// TIA Portal project "DistributoreCaffè" (V19) (continued)
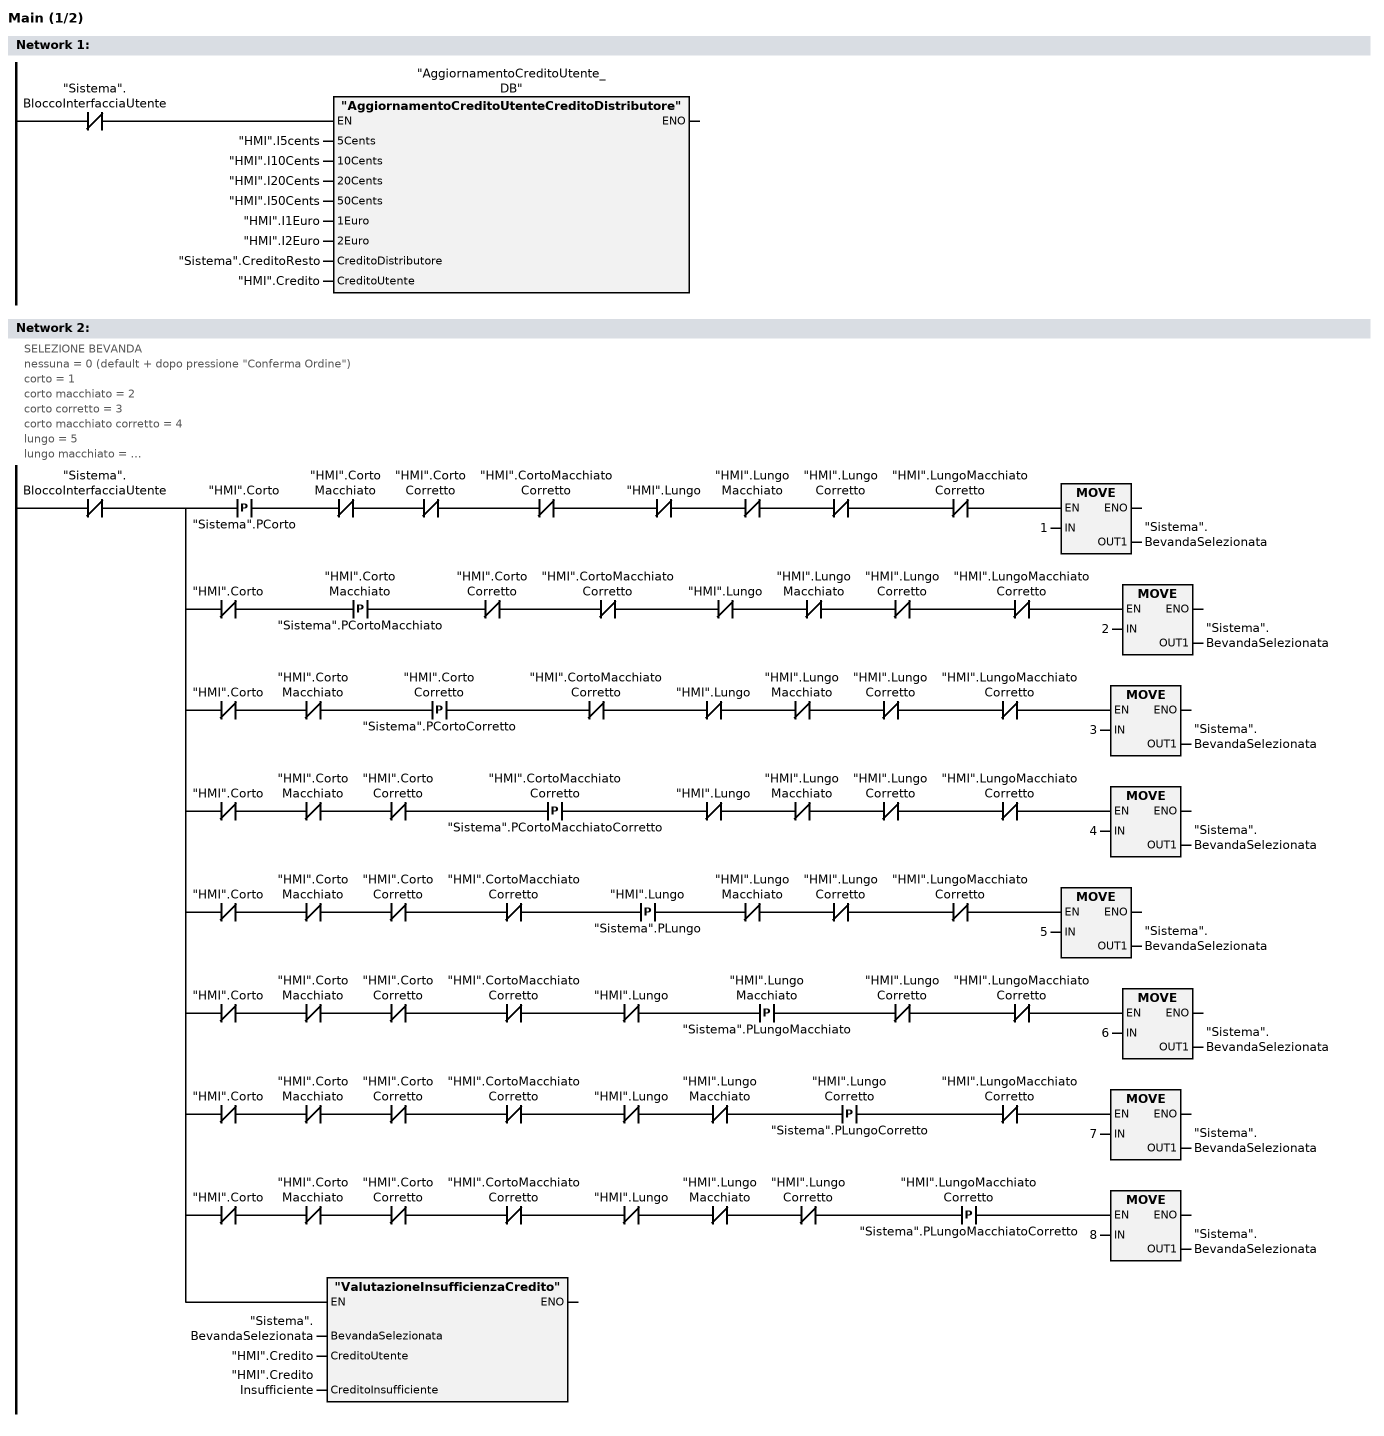
   RUNG wire#powerrail
      I_Contact( "Sistema".BloccoInterfacciaUtente )
      "AggiornamentoCreditoUtente_DB"("5Cents" := "HMI".I5cents, "10Cents" := "HMI".I10Cents, "20Cents" := "HMI".I20Cents, "50Cents" := "HMI".I50Cents, "1Euro" := "HMI".I1Euro, "2Euro" := "HMI".I2Euro, CreditoDistributore := "Sistema".CreditoResto, CreditoUtente := "HMI".Credito)
   END_RUNG
   // the same network as SCL:
   IF NOT "Sistema".BloccoInterfacciaUtente THEN
       "AggiornamentoCreditoUtente_DB"("5Cents" := "HMI".I5cents,   // "AggiornamentoCreditoUtenteCreditoDistributore"
                               "10Cents" := "HMI".I10Cents,
                               "20Cents" := "HMI".I20Cents,
                               "50Cents" := "HMI".I50Cents,
                               "1Euro" := "HMI".I1Euro,
                               "2Euro" := "HMI".I2Euro,
                               CreditoDistributore := "Sistema".CreditoResto,
                               CreditoUtente := "HMI".Credito);
   END_IF;
END_REGION

REGION Network 2
   // SELEZIONE BEVANDA
   // 
   // nessuna = 0 (default + dopo pressione "Conferma Ordine")
   // corto = 1
   // corto macchiato = 2
   // corto corretto = 3
   // corto macchiato corretto = 4
   // lungo = 5
   // lungo macchiato = 6
   // lungo corretto = 7
   // lungo macchiato corretto = 8
   // 
   // Il distributore avvisa con un lampeggio del diplay credito l'insufficienza di credito
   // 
   // Caso più pulsanti premuti contemporaneamente: priorità primo premuto
   RUNG wire#powerrail
      I_Contact( "Sistema".BloccoInterfacciaUtente )
      wire#w1
      P_Contact(operand := "HMI".Corto, bit := "Sistema".PCorto)
      I_Contact( "HMI".CortoMacchiato )
      I_Contact( "HMI".CortoCorretto )
      I_Contact( "HMI".CortoMacchiatoCorretto )
      I_Contact( "HMI".Lungo )
      I_Contact( "HMI".LungoMacchiato )
      I_Contact( "HMI".LungoCorretto )
      I_Contact( "HMI".LungoMacchiatoCorretto )
      Move(in := 1, out1 => "Sistema".BevandaSelezionata)
   END_RUNG
   RUNG wire#w1
      I_Contact( "HMI".Corto )
      P_Contact(operand := "HMI".CortoMacchiato, bit := "Sistema".PCortoMacchiato)
      I_Contact( "HMI".CortoCorretto )
      I_Contact( "HMI".CortoMacchiatoCorretto )
      I_Contact( "HMI".Lungo )
      I_Contact( "HMI".LungoMacchiato )
      I_Contact( "HMI".LungoCorretto )
      I_Contact( "HMI".LungoMacchiatoCorretto )
      Move(in := 2, out1 => "Sistema".BevandaSelezionata)
   END_RUNG
   RUNG wire#w1
      I_Contact( "HMI".Corto )
      I_Contact( "HMI".CortoMacchiato )
      P_Contact(operand := "HMI".CortoCorretto, bit := "Sistema".PCortoCorretto)
      I_Contact( "HMI".CortoMacchiatoCorretto )
      I_Contact( "HMI".Lungo )
      I_Contact( "HMI".LungoMacchiato )
      I_Contact( "HMI".LungoCorretto )
      I_Contact( "HMI".LungoMacchiatoCorretto )
      Move(in := 3, out1 => "Sistema".BevandaSelezionata)
   END_RUNG
   RUNG wire#w1
      I_Contact( "HMI".Corto )
      I_Contact( "HMI".CortoMacchiato )
      I_Contact( "HMI".CortoCorretto )
      P_Contact(operand := "HMI".CortoMacchiatoCorretto, bit := "Sistema".PCortoMacchiatoCorretto)
      I_Contact( "HMI".Lungo )
      I_Contact( "HMI".LungoMacchiato )
      I_Contact( "HMI".LungoCorretto )
      I_Contact( "HMI".LungoMacchiatoCorretto )
      Move(in := 4, out1 => "Sistema".BevandaSelezionata)
   END_RUNG
   RUNG wire#w1
      I_Contact( "HMI".Corto )
      I_Contact( "HMI".CortoMacchiato )
      I_Contact( "HMI".CortoCorretto )
      I_Contact( "HMI".CortoMacchiatoCorretto )
      P_Contact(operand := "HMI".Lungo, bit := "Sistema".PLungo)
      I_Contact( "HMI".LungoMacchiato )
      I_Contact( "HMI".LungoCorretto )
      I_Contact( "HMI".LungoMacchiatoCorretto )
      Move(in := 5, out1 => "Sistema".BevandaSelezionata)
   END_RUNG
   RUNG wire#w1
      I_Contact( "HMI".Corto )
      I_Contact( "HMI".CortoMacchiato )
      I_Contact( "HMI".CortoCorretto )
      I_Contact( "HMI".CortoMacchiatoCorretto )
      I_Contact( "HMI".Lungo )
      P_Contact(operand := "HMI".LungoMacchiato, bit := "Sistema".PLungoMacchiato)
      I_Contact( "HMI".LungoCorretto )
      I_Contact( "HMI".LungoMacchiatoCorretto )
      Move(in := 6, out1 => "Sistema".BevandaSelezionata)
   END_RUNG
   RUNG wire#w1
      I_Contact( "HMI".Corto )
      I_Contact( "HMI".CortoMacchiato )
      I_Contact( "HMI".CortoCorretto )
      I_Contact( "HMI".CortoMacchiatoCorretto )
      I_Contact( "HMI".Lungo )
      I_Contact( "HMI".LungoMacchiato )
      P_Contact(operand := "HMI".LungoCorretto, bit := "Sistema".PLungoCorretto)
      I_Contact( "HMI".LungoMacchiatoCorretto )
      Move(in := 7, out1 => "Sistema".BevandaSelezionata)
   END_RUNG
   RUNG wire#w1
      I_Contact( "HMI".Corto )
      I_Contact( "HMI".CortoMacchiato )
      I_Contact( "HMI".CortoCorretto )
      I_Contact( "HMI".CortoMacchiatoCorretto )
      I_Contact( "HMI".Lungo )
      I_Contact( "HMI".LungoMacchiato )
      I_Contact( "HMI".LungoCorretto )
      P_Contact(operand := "HMI".LungoMacchiatoCorretto, bit := "Sistema".PLungoMacchiatoCorretto)
      Move(in := 8, out1 => "Sistema".BevandaSelezionata)
   END_RUNG
   RUNG wire#w1
      "ValutazioneInsufficienzaCredito"(BevandaSelezionata := "Sistema".BevandaSelezionata, CreditoUtente := "HMI".Credito, CreditoInsufficiente := "HMI".CreditoInsufficiente)
   END_RUNG
   // the same network as SCL:
   #_w1 := NOT "Sistema".BloccoInterfacciaUtente;
   #_w2 := #_w1 AND "HMI".Corto AND NOT "Sistema".PCorto;   // rising edge of "HMI".Corto
   "Sistema".PCorto := "HMI".Corto;
   IF #_w2 AND NOT "HMI".CortoMacchiato AND NOT "HMI".CortoCorretto AND NOT "HMI".CortoMacchiatoCorretto AND NOT "HMI".Lungo AND NOT "HMI".LungoMacchiato AND NOT "HMI".LungoCorretto AND NOT "HMI".LungoMacchiatoCorretto THEN
       "Sistema".BevandaSelezionata := 1;
   END_IF;
   #_w3 := #_w1 AND NOT "HMI".Corto AND "HMI".CortoMacchiato AND NOT "Sistema".PCortoMacchiato;   // rising edge of "HMI".CortoMacchiato
   "Sistema".PCortoMacchiato := "HMI".CortoMacchiato;
   IF #_w3 AND NOT "HMI".CortoCorretto AND NOT "HMI".CortoMacchiatoCorretto AND NOT "HMI".Lungo AND NOT "HMI".LungoMacchiato AND NOT "HMI".LungoCorretto AND NOT "HMI".LungoMacchiatoCorretto THEN
       "Sistema".BevandaSelezionata := 2;
   END_IF;
   #_w4 := #_w1 AND NOT "HMI".Corto AND NOT "HMI".CortoMacchiato AND "HMI".CortoCorretto AND NOT "Sistema".PCortoCorretto;   // rising edge of "HMI".CortoCorretto
   "Sistema".PCortoCorretto := "HMI".CortoCorretto;
   IF #_w4 AND NOT "HMI".CortoMacchiatoCorretto AND NOT "HMI".Lungo AND NOT "HMI".LungoMacchiato AND NOT "HMI".LungoCorretto AND NOT "HMI".LungoMacchiatoCorretto THEN
       "Sistema".BevandaSelezionata := 3;
   END_IF;
   #_w5 := #_w1 AND NOT "HMI".Corto AND NOT "HMI".CortoMacchiato AND NOT "HMI".CortoCorretto AND "HMI".CortoMacchiatoCorretto AND NOT "Sistema".PCortoMacchiatoCorretto;   // rising edge of "HMI".CortoMacchiatoCorretto
   "Sistema".PCortoMacchiatoCorretto := "HMI".CortoMacchiatoCorretto;
   IF #_w5 AND NOT "HMI".Lungo AND NOT "HMI".LungoMacchiato AND NOT "HMI".LungoCorretto AND NOT "HMI".LungoMacchiatoCorretto THEN
       "Sistema".BevandaSelezionata := 4;
   END_IF;
   #_w6 := #_w1 AND NOT "HMI".Corto AND NOT "HMI".CortoMacchiato AND NOT "HMI".CortoCorretto AND NOT "HMI".CortoMacchiatoCorretto AND "HMI".Lungo AND NOT "Sistema".PLungo;   // rising edge of "HMI".Lungo
   "Sistema".PLungo := "HMI".Lungo;
   IF #_w6 AND NOT "HMI".LungoMacchiato AND NOT "HMI".LungoCorretto AND NOT "HMI".LungoMacchiatoCorretto THEN
       "Sistema".BevandaSelezionata := 5;
   END_IF;
   #_w7 := #_w1 AND NOT "HMI".Corto AND NOT "HMI".CortoMacchiato AND NOT "HMI".CortoCorretto AND NOT "HMI".CortoMacchiatoCorretto AND NOT "HMI".Lungo AND "HMI".LungoMacchiato AND NOT "Sistema".PLungoMacchiato;   // rising edge of "HMI".LungoMacchiato
   "Sistema".PLungoMacchiato := "HMI".LungoMacchiato;
   IF #_w7 AND NOT "HMI".LungoCorretto AND NOT "HMI".LungoMacchiatoCorretto THEN
       "Sistema".BevandaSelezionata := 6;
   END_IF;
   #_w8 := #_w1 AND NOT "HMI".Corto AND NOT "HMI".CortoMacchiato AND NOT "HMI".CortoCorretto AND NOT "HMI".CortoMacchiatoCorretto AND NOT "HMI".Lungo AND NOT "HMI".LungoMacchiato AND "HMI".LungoCorretto AND NOT "Sistema".PLungoCorretto;   // rising edge of "HMI".LungoCorretto
   "Sistema".PLungoCorretto := "HMI".LungoCorretto;
   IF #_w8 AND NOT "HMI".LungoMacchiatoCorretto THEN "Sistema".BevandaSelezionata := 7; END_IF;
   #_w9 := #_w1 AND NOT "HMI".Corto AND NOT "HMI".CortoMacchiato AND NOT "HMI".CortoCorretto AND NOT "HMI".CortoMacchiatoCorretto AND NOT "HMI".Lungo AND NOT "HMI".LungoMacchiato AND NOT "HMI".LungoCorretto AND "HMI".LungoMacchiatoCorretto AND NOT "Sistema".PLungoMacchiatoCorretto;   // rising edge of "HMI".LungoMacchiatoCorretto
   "Sistema".PLungoMacchiatoCorretto := "HMI".LungoMacchiatoCorretto;
   IF #_w9 THEN "Sistema".BevandaSelezionata := 8; END_IF;
   IF #_w1 THEN
       "ValutazioneInsufficienzaCredito"(BevandaSelezionata := "Sistema".BevandaSelezionata,
                               CreditoUtente := "HMI".Credito,
                               CreditoInsufficiente := "HMI".CreditoInsufficiente);
   END_IF;
END_REGION

REGION Network 3
   // Regolazione zucchero
   // 
   // Min = 0 unità
   // Max = 5 unità
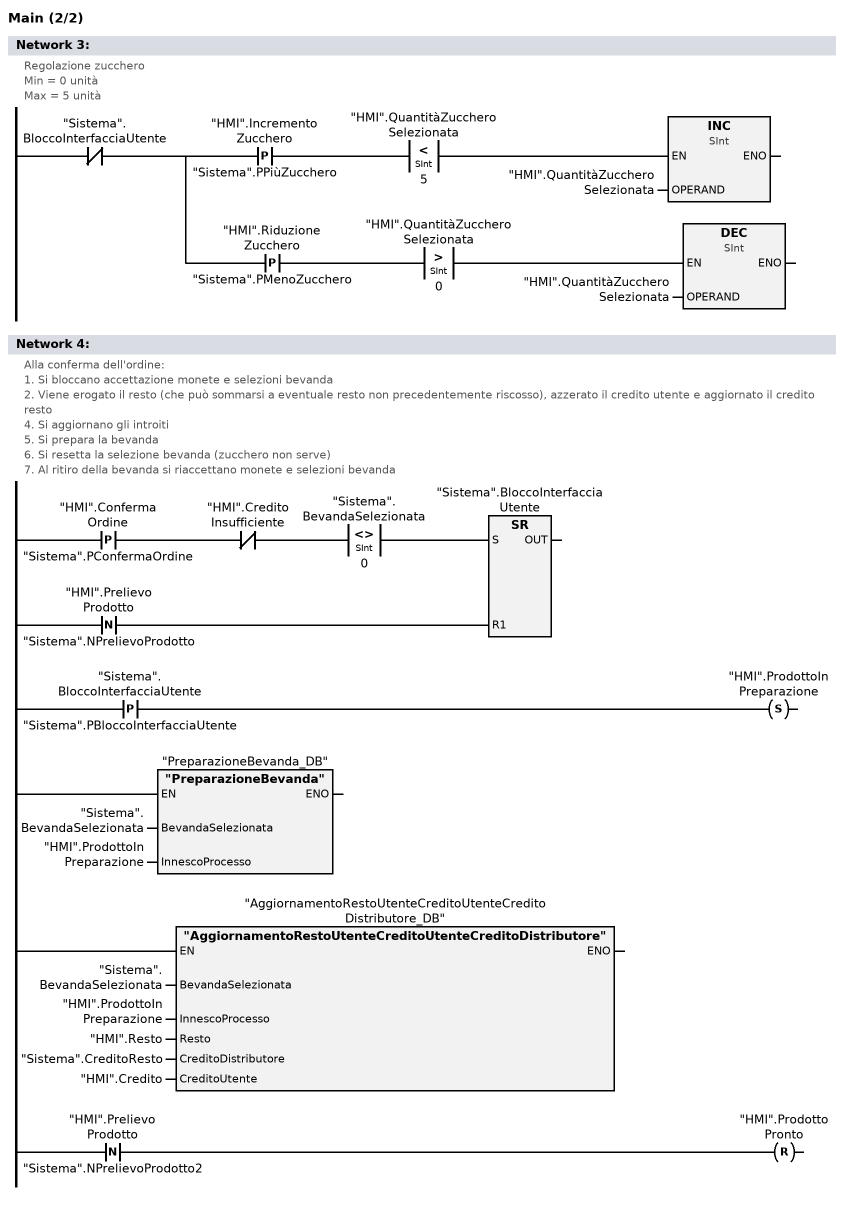
   RUNG wire#powerrail
      I_Contact( "Sistema".BloccoInterfacciaUtente )
      wire#w1
      P_Contact(operand := "HMI".IncrementoZucchero, bit := "Sistema".PPiùZucchero)
      { S7_Templates := "SrcType := SInt" } LT_Contact(in1 := "HMI".QuantitàZuccheroSelezionata, in2 := 5)
      { S7_Templates := "DestType := SInt" } Inc( "HMI".QuantitàZuccheroSelezionata )
   END_RUNG
   RUNG wire#w1
      P_Contact(operand := "HMI".RiduzioneZucchero, bit := "Sistema".PMenoZucchero)
      { S7_Templates := "SrcType := SInt" } GT_Contact(in1 := "HMI".QuantitàZuccheroSelezionata, in2 := 0)
      { S7_Templates := "DestType := SInt" } Dec( "HMI".QuantitàZuccheroSelezionata )
   END_RUNG
   // the same network as SCL:
   #_w1 := NOT "Sistema".BloccoInterfacciaUtente;
   #_w2 := #_w1 AND "HMI".IncrementoZucchero AND NOT "Sistema".PPiùZucchero;   // rising edge of "HMI".IncrementoZucchero
   "Sistema".PPiùZucchero := "HMI".IncrementoZucchero;
   IF #_w2 AND ("HMI".QuantitàZuccheroSelezionata < 5) THEN
       "HMI".QuantitàZuccheroSelezionata := "HMI".QuantitàZuccheroSelezionata + 1;
   END_IF;
   #_w3 := #_w1 AND "HMI".RiduzioneZucchero AND NOT "Sistema".PMenoZucchero;   // rising edge of "HMI".RiduzioneZucchero
   "Sistema".PMenoZucchero := "HMI".RiduzioneZucchero;
   IF #_w3 AND ("HMI".QuantitàZuccheroSelezionata > 0) THEN
       "HMI".QuantitàZuccheroSelezionata := "HMI".QuantitàZuccheroSelezionata - 1;
   END_IF;
END_REGION

REGION Network 4
   // Alla conferma dell'ordine:
   // 
   // 1. Si bloccano accettazione monete e selezioni bevanda
   // 2. Viene erogato il resto (che può sommarsi a eventuale resto non precedentemente riscosso), azzerato il credito utente e aggiornato il credito resto
   // 4. Si aggiornano gli introiti
   // 5. Si prepara la bevanda
   // 6. Si resetta la selezione bevanda (zucchero non serve)
   // 7. Al ritiro della bevanda si riaccettano monete e selezioni bevanda
   RUNG wire#powerrail
      P_Contact(operand := "HMI".ConfermaOrdine, bit := "Sistema".PConfermaOrdine)
      I_Contact( "HMI".CreditoInsufficiente )
      { S7_Templates := "SrcType := SInt" } NE_Contact(in1 := "Sistema".BevandaSelezionata, in2 := 0)
      S_SR(operand := "Sistema".BloccoInterfacciaUtente, r1 := wire#w1)
   END_RUNG
   RUNG wire#powerrail
      N_Contact(operand := "HMI".PrelievoProdotto, bit := "Sistema".NPrelievoProdotto)
   END_RUNG wire#w1
   RUNG wire#powerrail
      P_Contact(operand := "Sistema".BloccoInterfacciaUtente, bit := "Sistema".PBloccoInterfacciaUtente)
      S_Coil( "HMI".ProdottoInPreparazione )
   END_RUNG
   RUNG wire#powerrail
      "PreparazioneBevanda_DB"(BevandaSelezionata := "Sistema".BevandaSelezionata, InnescoProcesso := "HMI".ProdottoInPreparazione)
   END_RUNG
   RUNG wire#powerrail
      "AggiornamentoRestoUtenteCreditoUtenteCreditoDistributore_DB"(BevandaSelezionata := "Sistema".BevandaSelezionata, InnescoProcesso := "HMI".ProdottoInPreparazione, Resto := "HMI".Resto, CreditoDistributore := "Sistema".CreditoResto, CreditoUtente := "HMI".Credito)
   END_RUNG
   RUNG wire#powerrail
      N_Contact(operand := "HMI".PrelievoProdotto, bit := "Sistema".NPrelievoProdotto2)
      R_Coil( "HMI".ProdottoPronto )
   END_RUNG
   // the same network as SCL:
   #_w1 := "HMI".ConfermaOrdine AND NOT "Sistema".PConfermaOrdine;   // rising edge of "HMI".ConfermaOrdine
   "Sistema".PConfermaOrdine := "HMI".ConfermaOrdine;
   #_w2 := NOT "HMI".PrelievoProdotto AND "Sistema".NPrelievoProdotto;   // falling edge of "HMI".PrelievoProdotto
   "Sistema".NPrelievoProdotto := "HMI".PrelievoProdotto;
   IF #_w1 AND NOT "HMI".CreditoInsufficiente AND ("Sistema".BevandaSelezionata <> 0) THEN
       "Sistema".BloccoInterfacciaUtente := TRUE;   // SR flip-flop
   END_IF;
   IF #_w2 THEN "Sistema".BloccoInterfacciaUtente := FALSE; END_IF;
   #_w3 := "Sistema".BloccoInterfacciaUtente AND NOT "Sistema".PBloccoInterfacciaUtente;   // rising edge of "Sistema".BloccoInterfacciaUtente
   "Sistema".PBloccoInterfacciaUtente := "Sistema".BloccoInterfacciaUtente;
   IF #_w3 THEN "HMI".ProdottoInPreparazione := TRUE; END_IF;
   "PreparazioneBevanda_DB"(BevandaSelezionata := "Sistema".BevandaSelezionata,   // "PreparazioneBevanda"
                           InnescoProcesso := "HMI".ProdottoInPreparazione);
   "AggiornamentoRestoUtenteCreditoUtenteCreditoDistributore_DB"(BevandaSelezionata := "Sistema".BevandaSelezionata,   // "AggiornamentoRestoUtenteCreditoUtenteCreditoDistributore"
                           InnescoProcesso := "HMI".ProdottoInPreparazione,
                           Resto := "HMI".Resto,
                           CreditoDistributore := "Sistema".CreditoResto,
                           CreditoUtente := "HMI".Credito);
   #_w4 := NOT "HMI".PrelievoProdotto AND "Sistema".NPrelievoProdotto2;   // falling edge of "HMI".PrelievoProdotto
   "Sistema".NPrelievoProdotto2 := "HMI".PrelievoProdotto;
   IF #_w4 THEN "HMI".ProdottoPronto := FALSE; END_IF;
END_REGION
END_ORGANIZATION_BLOCK

(* ===== HMI "HMI_RT_1" =====
system functions are stored by id; their names below are inferred from use
connection "HMI_Collegamento_1": ETHERNET, SMART_S7_1200_OMS

HMI tags "Tabella delle variabili standard"
   "Variabile_Numero di pagina" : UInt, internal
   "HMI_ProdottoPronto" : Bool = PLC HMI.ProdottoPronto, 100 ms
   "HMI_PrelievoProdotto" : Bool = PLC HMI.PrelievoProdotto, 100 ms
   "HMI_BicchieriScarico" : Bool = PLC HMI.BicchieriScarico, 100 ms
   "HMI_PaletteScarico" : Bool = PLC HMI.PaletteScarico, 100 ms
   "HMI_CaffèScarico" : Bool = PLC HMI.CaffèScarico, 100 ms
   "HMI_LatteScarico" : Bool = PLC HMI.LatteScarico, 100 ms
   "HMI_GrappaScarico" : Bool = PLC HMI.GrappaScarico, 100 ms
   "HMI_ZuccheroScarico" : Bool = PLC HMI.ZuccheroScarico, 100 ms
   "HMI_Bicchieri" : Int = PLC HMI.Bicchieri, 100 ms
   "HMI_Palette" : Int = PLC HMI.Palette, 100 ms
   "HMI_Caffè" : SInt = PLC HMI.Caffè, 100 ms
   "HMI_Latte" : SInt = PLC HMI.Latte, 100 ms
   "HMI_Grappa" : SInt = PLC HMI.Grappa, 100 ms
   "HMI_Zucchero" : SInt = PLC HMI.Zucchero, 100 ms
   "HMI_Credito" : Real = PLC HMI.Credito, 100 ms
   "HMI_Introiti" : Real = PLC HMI.Introiti, 100 ms
   "HMI_PrelievoIntroiti" : Bool = PLC HMI.PrelievoIntroiti, 100 ms
   "HMI_CreditoInsufficiente" : Bool = PLC HMI.CreditoInsufficiente, 100 ms
   "HMI_I5cents" : Bool = PLC HMI.I5cents, 100 ms
   "HMI_I10Cents" : Bool = PLC HMI.I10Cents, 100 ms
   "HMI_I20Cents" : Bool = PLC HMI.I20Cents, 100 ms
   "HMI_I50Cents" : Bool = PLC HMI.I50Cents, 100 ms
   "HMI_I1Euro" : Bool = PLC HMI.I1Euro, 100 ms
   "HMI_I2Euro" : Bool = PLC HMI.I2Euro, 100 ms
   "HMI_Corto" : Bool = PLC HMI.Corto, 100 ms
   "HMI_CortoMacchiato" : Bool = PLC HMI.CortoMacchiato, 100 ms
   "HMI_CortoCorretto" : Bool = PLC HMI.CortoCorretto, 100 ms
   "HMI_CortoMacchiatoCorretto" : Bool = PLC HMI.CortoMacchiatoCorretto, 100 ms
   "HMI_Lungo" : Bool = PLC HMI.Lungo, 100 ms
   "HMI_LungoMacchiato" : Bool = PLC HMI.LungoMacchiato, 100 ms
   "HMI_LungoCorretto" : Bool = PLC HMI.LungoCorretto, 100 ms
   "HMI_LungoMacchiatoCorretto" : Bool = PLC HMI.LungoMacchiatoCorretto, 100 ms
   "HMI_ValvolaBicchiere" : Bool = PLC HMI.ValvolaBicchiere, 100 ms
   "HMI_ValvolaZucchero" : Bool = PLC HMI.ValvolaZucchero, 100 ms
   "HMI_ValvolaGrappa" : Bool = PLC HMI.ValvolaGrappa, 100 ms
   "HMI_ValvolaLatte" : Bool = PLC HMI.ValvolaLatte, 100 ms
   "HMI_ValvolaCaffè" : Bool = PLC HMI.ValvolaCaffè, 100 ms
   "HMI_ValvolaPaletta" : Bool = PLC HMI.ValvolaPaletta, 100 ms
   "HMI_QuantitàZuccheroSelezionata" : SInt = PLC HMI.QuantitàZuccheroSelezionata, 100 ms
   "HMI_RiduzioneZucchero" : Bool = PLC HMI.RiduzioneZucchero, 100 ms
   "HMI_IncrementoZucchero" : Bool = PLC HMI.IncrementoZucchero, 100 ms
   "HMI_ConfermaOrdine" : Bool = PLC HMI.ConfermaOrdine, 100 ms
   "HMI_Resto" : RestoUtente = PLC HMI.Resto, 100 ms
   "HMI_Resto_5Cents" : SInt = PLC HMI.Resto.5Cents, 100 ms
   "HMI_Resto_10Cents" : SInt = PLC HMI.Resto.10Cents, 100 ms
   "HMI_Resto_20Cents" : SInt = PLC HMI.Resto.20Cents, 100 ms
   "HMI_Resto_50Cents" : SInt = PLC HMI.Resto.50Cents, 100 ms
   "HMI_Resto_1Euro" : SInt = PLC HMI.Resto.1Euro, 100 ms
   "HMI_Resto_2Euro" : SInt = PLC HMI.Resto.2Euro, 100 ms
   "HMI_ProdottoInPreparazione" : Bool = PLC HMI.ProdottoInPreparazione, 100 ms

text list "Elenco testi_Nome della pagina": 1 'Pagina base'; 2 'Gestione utenti'

Template "Modello_1" 800x480
   Button "Pagina iniziale" at 1,39 size 55x39; TextOff 'Pagina iniziale'; PictureOff "NavigateHome_KTP900_Basic_PN_TR"; PictureOn "NavigateHome_KTP900_Basic_PN_TR"
      on Release: ActivateScreen("Distributore", 0)
   Button "Template_Button" at 1,79 size 55x39; TextOff 'Text'
   Button "Template_Button_1" at 1,119 size 55x39; TextOff 'Text'
   Button "Template_Button_2" at 1,159 size 55x39; TextOff 'Text'
   Button "Template_Button_3" at 1,199 size 55x39; TextOff 'Text'
   Button "Template_Button_4" at 1,239 size 55x39; TextOff 'Text'
   Button "Template_Button_5" at 1,279 size 55x39; TextOff 'Text'
   Button "Template_Button_6" at 1,319 size 55x39; TextOff 'Text'
   Button "Template_Button_7" at 1,359 size 55x39; TextOff 'Text'
   Button "Connessione" at 1,399 size 55x39; TextOff 'Connessione'; PictureOff "Login_KTP900_Basic_PN_TR"; PictureOn "Login_KTP900_Basic_PN_TR"
      on Release: function_a2a04561()
   Button "Esci" at 1,439 size 55x39; TextOff 'Esci'; PictureOff "ExitRuntime_KTP900_Basic_PN_TR"; PictureOn "ExitRuntime_KTP900_Basic_PN_TR"
      on Release: StopRuntime(0)
   SymbolicIOField "Pagina_campo_IO_simbolico" at 2,7 size 691x26; TextOff '0'; TextOn '1'; TextList "Elenco testi_Nome della pagina"
      ProcessValue <- "Variabile_Numero di pagina"
      on Change: ActivateScreenByNumber("Variabile_Numero di pagina", 0)
   DateTimeField "HmiScreenItemData" at 695,20 size 105x20
   DateTimeField "HmiScreenItemData_1" at 695,0 size 105x20

screen "Distributore" 800x480, template "Modello_1"
   on GenerateScreen: SetTag("Variabile_Numero di pagina", 1)
   Button "Pulsante_1" at 77,61 size 96x32; TextOff '0,05€'; TextOn '0,05'
      on Press: SetBit("HMI_I5cents")
      on Release: ResetBit("HMI_I5cents")
   TextField "Casella di testo_1" at 59,39 size 133x20; Text 'Inserimento credito'
   Button "Pulsante_2" at 77,93 size 96x32; TextOff '0,10€'; TextOn '0,10'
      on Press: SetBit("HMI_I10Cents")
      on Release: ResetBit("HMI_I10Cents")
   Button "Pulsante_3" at 77,125 size 96x32; TextOff '0,20€'; TextOn '0,20'
      on Press: SetBit("HMI_I20Cents")
      on Release: ResetBit("HMI_I20Cents")
   Button "Pulsante_4" at 77,157 size 96x32; TextOff '0,50€'; TextOn '0,50'
      on Press: SetBit("HMI_I50Cents")
      on Release: ResetBit("HMI_I50Cents")
   Button "Pulsante_5" at 77,189 size 96x32; TextOff '1€'; TextOn '1'
      on Press: SetBit("HMI_I1Euro")
      on Release: ResetBit("HMI_I1Euro")
   Button "Pulsante_6" at 77,221 size 96x32; TextOff '2€'; TextOn '2'
      on Press: SetBit("HMI_I2Euro")
      on Release: ResetBit("HMI_I2Euro")
   TextField "Casella di testo_2" at 310,41 size 96x20; Text 'Prelievo resto'
   Button "Pulsante_7" at 292,66 size 60x60; TextOff 'Text'; PictureOff "5cents"; PictureOn "5cents"
      on Click: function_b9b71300("HMI_Resto_5Cents", 1)
      Visibility <- "HMI_Resto_5Cents"
   Button "Pulsante_8" at 368,66 size 60x60; TextOff 'Text'; PictureOff "10cents"; PictureOn "10cents"
      on Click: function_b9b71300("HMI_Resto_10Cents", 1)
      Visibility <- "HMI_Resto_10Cents"
   Button "Pulsante_9" at 292,134 size 60x60; TextOff 'Text'; PictureOff "20cents"; PictureOn "20cents"
      on Click: function_b9b71300("HMI_Resto_20Cents", 1)
      Visibility <- "HMI_Resto_20Cents"
   Button "Pulsante_10" at 368,134 size 60x60; TextOff 'Text'; PictureOff "50cents"; PictureOn "50cents"
      on Click: function_b9b71300("HMI_Resto_50Cents", 1)
      Visibility <- "HMI_Resto_50Cents"
   Button "Pulsante_11" at 292,204 size 60x60; TextOff 'Text'; PictureOff "1euro"; PictureOn "1euro"
      on Click: function_b9b71300("HMI_Resto_1Euro", 1)
      Visibility <- "HMI_Resto_1Euro"
   Button "Pulsante_12" at 368,204 size 60x60; TextOff 'Text'; PictureOff "2euro"; PictureOn "2euro"
      on Click: function_b9b71300("HMI_Resto_2Euro", 1)
      Visibility <- "HMI_Resto_2Euro"
   IOField "Campo I/O_1" at 245,83 size 37x32; FormatPattern 99
      ProcessValue <- "HMI_Resto_5Cents"
   IOField "Campo I/O_2" at 245,147 size 37x32; FormatPattern 99
      ProcessValue <- "HMI_Resto_20Cents"
   IOField "Campo I/O_3" at 245,216 size 37x32; FormatPattern 99
      ProcessValue <- "HMI_Resto_1Euro"
   IOField "Campo I/O_4" at 440,83 size 37x32; FormatPattern 99
      ProcessValue <- "HMI_Resto_10Cents"
   IOField "Campo I/O_5" at 440,147 size 37x32; FormatPattern 99
      ProcessValue <- "HMI_Resto_50Cents"
   IOField "Campo I/O_6" at 440,216 size 37x32; FormatPattern 99
      ProcessValue <- "HMI_Resto_2Euro"
   IOField "Campo I/O_7" at 100,278 size 49x32; FormatPattern 99.99
      ProcessValue <- "HMI_Credito"
      Appearance <- "HMI_CreditoInsufficiente"
   TextField "Casella di testo_3" at 96,257 size 52x20; Text 'Credito'
   Group "Group" at 566,286 size 89x83; Picture "Grafica_6"
   Group "Group_1" at 566,174 size 89x83; Picture "Grafica_6"
   Group "Group_3" at 701,286 size 89x83; Picture "Grafica_6"
   Group "Group_4" at 701,174 size 89x83; Picture "Grafica_6"
   Group "Group_5" at 701,64 size 89x83; Picture "Grafica_6"
   TextField "Casella di testo_5" at 701,43 size 52x20; Text 'Paletta'
   TextField "Casella di testo_6" at 572,152 size 39x20; Text 'Caffè'
   TextField "Casella di testo_7" at 707,154 size 40x20; Text 'Latte'
   TextField "Casella di testo_8" at 566,266 size 51x20; Text 'Grappa'
   TextField "Casella di testo_9" at 695,266 size 64x20; Text 'Zucchero'
   Group "Group_6" at 562,44 size 93x103; Picture "Grafica_6"
   Button "Pulsante_13" at 617,372 size 82x82; TextOff 'Text'; PictureOff "BevandaPronta"; PictureOn "BevandaPronta_1"
      Visibility <- "HMI_ProdottoPronto"
      on Press: SetBit("HMI_PrelievoProdotto")
      on Release: ResetBit("HMI_PrelievoProdotto")
   GraphicView "Vista grafica_19" at 588,375 size 145x76; Picture "PaoloBitta"
      Visibility <- "HMI_ProdottoInPreparazione"
   TextField "Casella di testo_10" at 322,300 size 126x20; Text 'Selezione bevanda'
   Button "Pulsante_14" at 207,323 size 175x32; TextOff 'Corto 0,30€'; TextOn 'Corto'
      on Press: SetBit("HMI_Corto")
      on Release: ResetBit("HMI_Corto")
   Button "Pulsante_15" at 382,323 size 175x32; TextOff 'Corto macchiato 0,40€'; TextOn 'Corto macchiato'
      on Press: SetBit("HMI_CortoMacchiato")
      on Release: ResetBit("HMI_CortoMacchiato")
   Button "Pulsante_16" at 382,355 size 175x32; TextOff 'Corto corretto 0,40€'; TextOn 'Corto corretto'
      on Press: SetBit("HMI_CortoCorretto")
      on Release: ResetBit("HMI_CortoCorretto")
   Button "Pulsante_17" at 207,355 size 175x32; TextOff 'Corto macchiato corretto 0,50€'; TextOn 'Corto macchiato corretto'
      on Press: SetBit("HMI_CortoMacchiatoCorretto")
      on Release: ResetBit("HMI_CortoMacchiatoCorretto")
   Button "Pulsante_18" at 207,391 size 175x32; TextOff 'Lungo 0,60€'; TextOn 'Lungo'
      on Press: SetBit("HMI_Lungo")
      on Release: ResetBit("HMI_Lungo")
   Button "Pulsante_19" at 382,391 size 175x32; TextOff 'Lungo macchiato 0,70€'; TextOn 'Lungo macchiato'
      on Release: ResetBit("HMI_LungoMacchiato")
      on Press: SetBit("HMI_LungoMacchiato")
   Button "Pulsante_20" at 382,423 size 175x32; TextOff 'Lungo corretto 0,70€'; TextOn 'Lungo corretto'
      on Press: SetBit("HMI_LungoCorretto")
      on Release: ResetBit("HMI_LungoCorretto")
   Button "Pulsante_21" at 207,423 size 175x32; TextOff 'Lungo macchiato corretto 0,80€'; TextOn 'Lungo macchiato corretto'
      on Press: SetBit("HMI_LungoMacchiatoCorretto")
      on Release: ResetBit("HMI_LungoMacchiatoCorretto")
   TextField "Casella di testo_11" at 59,328 size 146x20; Text 'Regolazione zucchero'
   Button "Pulsante_22" at 65,355 size 38x32; TextOff '-'
      on Press: SetBit("HMI_RiduzioneZucchero")
      on Release: ResetBit("HMI_RiduzioneZucchero")
   Button "Pulsante_23" at 161,355 size 37x32; TextOff '+'
      on Release: ResetBit("HMI_IncrementoZucchero")
      on Press: SetBit("HMI_IncrementoZucchero")
   IOField "Campo I/O_8" at 114,355 size 36x32; FormatPattern 9
      ProcessValue <- "HMI_QuantitàZuccheroSelezionata"
   Button "Pulsante_24" at 73,422 size 119x32; TextOff 'Conferma ordine'
      on Press: SetBit("HMI_ConfermaOrdine")
      on Release: ResetBit("HMI_ConfermaOrdine")
   GraphicView "Vista grafica_10" at 566,286 size 69x83; Picture "Grafica_6"
   GraphicView "Vista grafica_9" at 622,306 size 19x43; Picture "Grafica_5"
      Visibility <- "HMI_ValvolaGrappa"
   GraphicView "Vista grafica_8" at 608,316 size 47x23; Picture "Grafica_4"
      Visibility <- "HMI_ValvolaGrappa"
   GraphicView "Vista grafica_1" at 566,174 size 69x83; Picture "Grafica_6"
   GraphicView "Vista grafica_2" at 622,194 size 19x43; Picture "Grafica_5"
      Visibility <- "HMI_ValvolaCaffè"
   GraphicView "Vista grafica_3" at 608,204 size 47x23; Picture "Grafica_4"
      Visibility <- "HMI_ValvolaCaffè"
   GraphicView "Vista grafica_4" at 566,64 size 69x83; Picture "Grafica_6"
   GraphicView "Vista grafica_5" at 622,84 size 19x43; Picture "Grafica_5"
      Visibility <- "HMI_ValvolaBicchiere"
   GraphicView "Vista grafica_6" at 608,94 size 47x23; Picture "Grafica_4"
      Visibility <- "HMI_ValvolaBicchiere"
   Group "Group_2" at 566,64 size 89x83; Picture "Grafica_6"
   TextField "Casella di testo_4" at 562,44 size 63x20; Text 'Bicchiere'
   GraphicView "Vista grafica_7" at 701,286 size 69x83; Picture "Grafica_6"
   GraphicView "Vista grafica_11" at 757,306 size 19x43; Picture "Grafica_5"
      Visibility <- "HMI_ValvolaZucchero"
   GraphicView "Vista grafica_12" at 743,316 size 47x23; Picture "Grafica_4"
      Visibility <- "HMI_ValvolaZucchero"
   GraphicView "Vista grafica_13" at 701,174 size 69x83; Picture "Grafica_6"
   GraphicView "Vista grafica_14" at 757,194 size 19x43; Picture "Grafica_5"
      Visibility <- "HMI_ValvolaLatte"
   GraphicView "Vista grafica_15" at 743,204 size 47x23; Picture "Grafica_4"
      Visibility <- "HMI_ValvolaLatte"
   GraphicView "Vista grafica_16" at 701,64 size 69x83; Picture "Grafica_6"
   GraphicView "Vista grafica_17" at 757,84 size 19x43; Picture "Grafica_5"
      Visibility <- "HMI_ValvolaPaletta"
   GraphicView "Vista grafica_18" at 743,94 size 47x23; Picture "Grafica_4"
      Visibility <- "HMI_ValvolaPaletta"

screen "Gestione utenti" 800x480, template "Modello_1"
   on GenerateScreen: SetTag("Variabile_Numero di pagina", 2)
   UserView "HmiScreenItemData" at 57,89 size 740x383
   Button "Indietro" at 57,41 size 159x47; TextOff 'Indietro'
      on Release: ActivateScreen("Distributore", 0)

screen "Serbatoi" 800x480
   Bar "Barra grafica_1" at 647,86 size 100x200; MinimumValue 0; MaximumValue 100
      ProcessValue <- "HMI_Zucchero"
   Bar "Barra grafica_2" at 498,85 size 100x200; MinimumValue 0; MaximumValue 100
      ProcessValue <- "HMI_Grappa"
   Bar "Barra grafica_3" at 357,84 size 100x200; MinimumValue 0; MaximumValue 100
      ProcessValue <- "HMI_Latte"
   Bar "Barra grafica_4" at 234,84 size 100x200; MinimumValue 0; MaximumValue 100
      ProcessValue <- "HMI_Caffè"
   IOField "Campo I/O_1" at 90,108 size 96x32; FormatPattern 99999
      ProcessValue <- "HMI_Bicchieri"
   IOField "Campo I/O_2" at 87,200 size 96x32; FormatPattern 99999
      ProcessValue <- "HMI_Palette"
   TextField "Casella di testo_1" at 106,84 size 58x20; Text 'Bicchieri'
   TextField "Casella di testo_2" at 105,178 size 52x20; Text 'Palette'
   TextField "Casella di testo_3" at 262,58 size 39x20; Text 'Caffè'
   TextField "Casella di testo_4" at 387,58 size 40x20; Text 'Latte'
   TextField "Casella di testo_5" at 524,58 size 51x20; Text 'Grappa'
   TextField "Casella di testo_6" at 668,58 size 64x20; Text 'Zucchero'
   GraphicIOField "PlotLight_Square_N_Mono" at 21,92 size 50x50; PictureOff "PilotLight_Square_N_Off_mono"; PictureOn "PilotLight_Square_N_On_mono"
      ProcessValue <- "HMI_BicchieriScarico"
      Appearance <- "HMI_BicchieriScarico"
   GraphicIOField "PlotLight_Square_N_Mono_1" at 259,293 size 50x50; PictureOff "PilotLight_Square_N_Off_mono"; PictureOn "PilotLight_Square_N_On_mono"
      ProcessValue <- "HMI_CaffèScarico"
      Appearance <- "HMI_CaffèScarico"
   GraphicIOField "PlotLight_Square_N_Mono_2" at 387,293 size 50x50; PictureOff "PilotLight_Square_N_Off_mono"; PictureOn "PilotLight_Square_N_On_mono"
      Appearance <- "HMI_LatteScarico"
      ProcessValue <- "HMI_LatteScarico"
   GraphicIOField "PlotLight_Square_N_Mono_3" at 521,292 size 50x50; PictureOff "PilotLight_Square_N_Off_mono"; PictureOn "PilotLight_Square_N_On_mono"
      ProcessValue <- "HMI_GrappaScarico"
      Appearance <- "HMI_GrappaScarico"
   GraphicIOField "PlotLight_Square_N_Mono_4" at 675,292 size 50x50; PictureOff "PilotLight_Square_N_Off_mono"; PictureOn "PilotLight_Square_N_On_mono"
      Appearance <- "HMI_ZuccheroScarico"
      ProcessValue <- "HMI_ZuccheroScarico"
   GraphicIOField "PlotLight_Square_N_Mono_5" at 19,186 size 50x50; PictureOff "PilotLight_Square_N_Off_mono"; PictureOn "PilotLight_Square_N_On_mono"
      ProcessValue <- "HMI_PaletteScarico"
      Appearance <- "HMI_PaletteScarico"

screen "InfoAdmin" 800x480
   TextField "Casella di testo_1" at 64,27 size 50x20; Text 'Introiti'
   IOField "Campo I/O_1" at 37,52 size 108x32; FormatPattern 999.99
      ProcessValue <- "HMI_Introiti"
   Button "Pulsante_1" at 159,52 size 96x32; TextOff 'Prelievo'
      on Press: SetBit("HMI_PrelievoIntroiti")
      on Release: ResetBit("HMI_PrelievoIntroiti")
*)